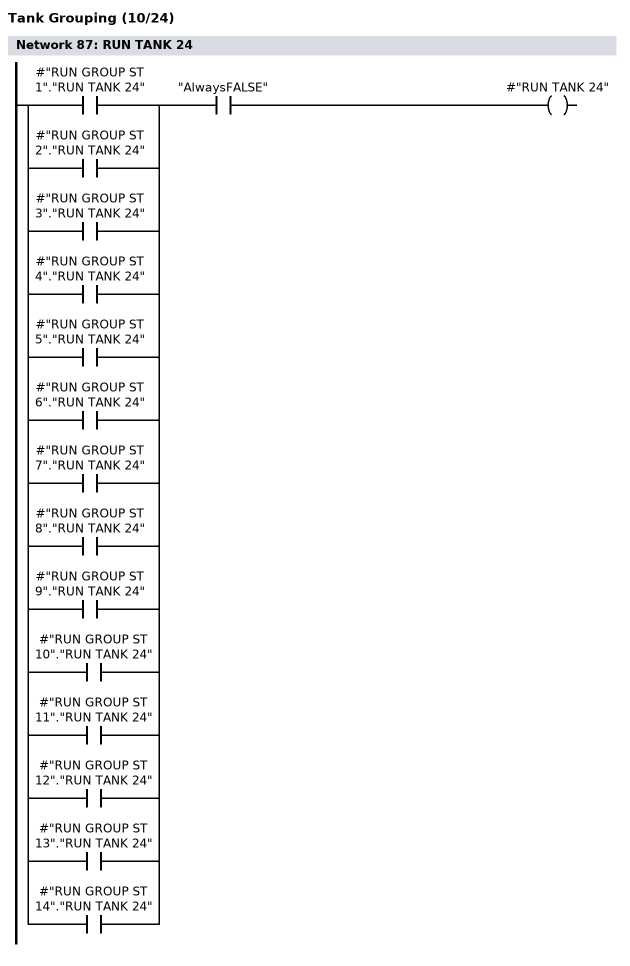
   RUNG wire#powerrail
      Contact( #"RUN GROUP ST 1"."RUN TANK 24" )
      wire#w1
      Contact( "AlwaysFALSE" )
      Coil( #"RUN TANK 24" )
   END_RUNG
   RUNG wire#powerrail
      Contact( #"RUN GROUP ST 2"."RUN TANK 24" )
   END_RUNG wire#w1
   RUNG wire#powerrail
      Contact( #"RUN GROUP ST 3"."RUN TANK 24" )
   END_RUNG wire#w1
   RUNG wire#powerrail
      Contact( #"RUN GROUP ST 4"."RUN TANK 24" )
   END_RUNG wire#w1
   RUNG wire#powerrail
      Contact( #"RUN GROUP ST 5"."RUN TANK 24" )
   END_RUNG wire#w1
   RUNG wire#powerrail
      Contact( #"RUN GROUP ST 6"."RUN TANK 24" )
   END_RUNG wire#w1
   RUNG wire#powerrail
      Contact( #"RUN GROUP ST 7"."RUN TANK 24" )
   END_RUNG wire#w1
   RUNG wire#powerrail
      Contact( #"RUN GROUP ST 8"."RUN TANK 24" )
   END_RUNG wire#w1
   RUNG wire#powerrail
      Contact( #"RUN GROUP ST 9"."RUN TANK 24" )
   END_RUNG wire#w1
   RUNG wire#powerrail
      Contact( #"RUN GROUP ST 10"."RUN TANK 24" )
   END_RUNG wire#w1
   RUNG wire#powerrail
      Contact( #"RUN GROUP ST 11"."RUN TANK 24" )
   END_RUNG wire#w1
   RUNG wire#powerrail
      Contact( #"RUN GROUP ST 12"."RUN TANK 24" )
   END_RUNG wire#w1
   RUNG wire#powerrail
      Contact( #"RUN GROUP ST 13"."RUN TANK 24" )
   END_RUNG wire#w1
   RUNG wire#powerrail
      Contact( #"RUN GROUP ST 14"."RUN TANK 24" )
   END_RUNG wire#w1
   // the same network as SCL:
   #"RUN TANK 24" := (#"RUN GROUP ST 1"."RUN TANK 24" OR #"RUN GROUP ST 2"."RUN TANK 24" OR #"RUN GROUP ST 3"."RUN TANK 24" OR #"RUN GROUP ST 4"."RUN TANK 24" OR #"RUN GROUP ST 5"."RUN TANK 24" OR #"RUN GROUP ST 6"."RUN TANK 24" OR #"RUN GROUP ST 7"."RUN TANK 24" OR #"RUN GROUP ST 8"."RUN TANK 24" OR #"RUN GROUP ST 9"."RUN TANK 24" OR #"RUN GROUP ST 10"."RUN TANK 24" OR #"RUN GROUP ST 11"."RUN TANK 24" OR #"RUN GROUP ST 12"."RUN TANK 24" OR #"RUN GROUP ST 13"."RUN TANK 24" OR #"RUN GROUP ST 14"."RUN TANK 24") AND "AlwaysFALSE";
END_REGION

REGION Network 89: Tank Selected Group 1
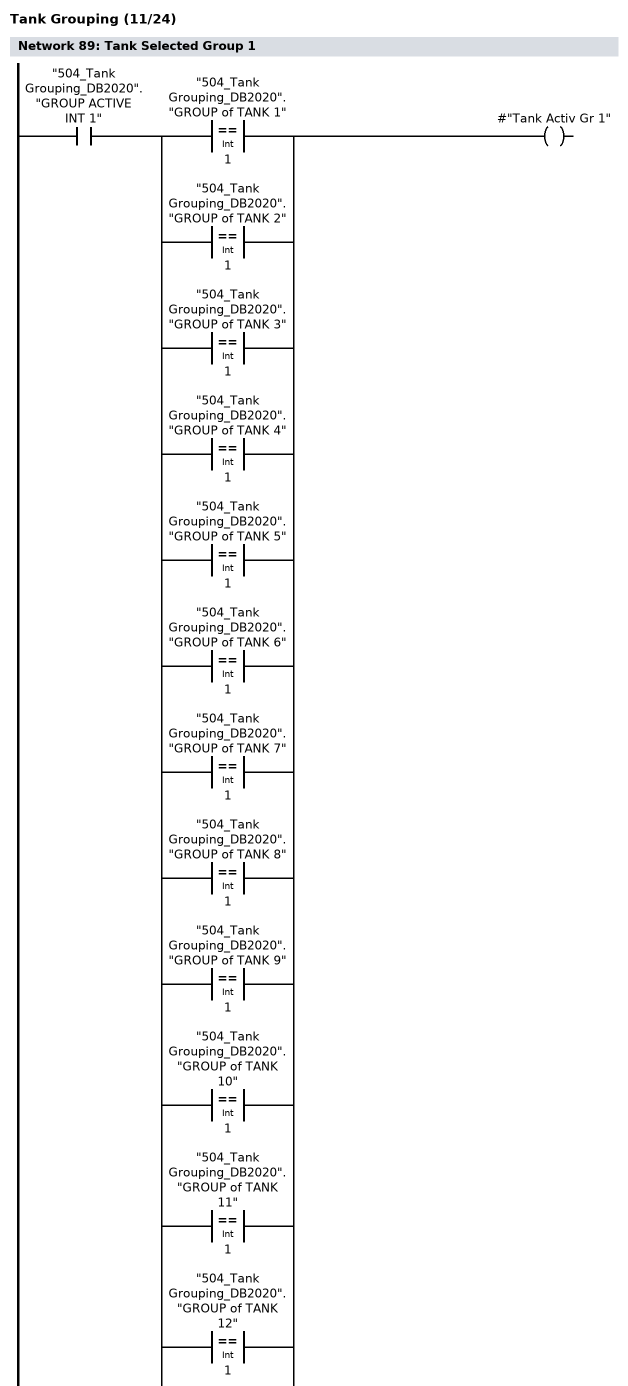
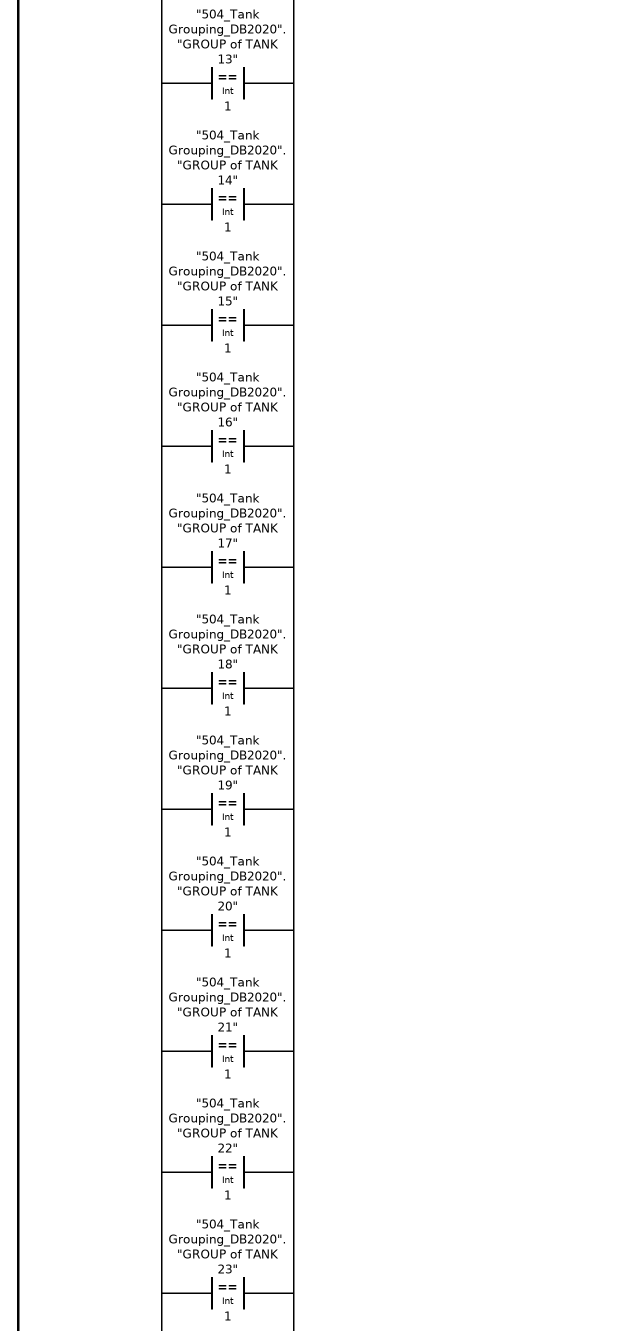
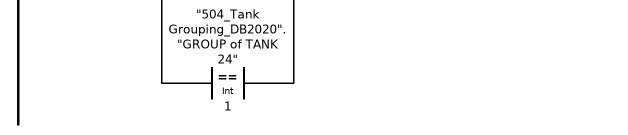
   RUNG wire#powerrail
      Contact( "504_Tank Grouping_DB2020"."GROUP ACTIVE INT 1" )
      wire#w1
      { S7_Templates := "SrcType := Int" } EQ_Contact(in1 := "504_Tank Grouping_DB2020"."GROUP of TANK 1", in2 := 1)
      wire#w2
      Coil( #"Tank Activ Gr 1" )
   END_RUNG
   RUNG wire#w1
      { S7_Templates := "SrcType := Int" } EQ_Contact(in1 := "504_Tank Grouping_DB2020"."GROUP of TANK 2", in2 := 1)
   END_RUNG wire#w2
   RUNG wire#w1
      { S7_Templates := "SrcType := Int" } EQ_Contact(in1 := "504_Tank Grouping_DB2020"."GROUP of TANK 3", in2 := 1)
   END_RUNG wire#w2
   RUNG wire#w1
      { S7_Templates := "SrcType := Int" } EQ_Contact(in1 := "504_Tank Grouping_DB2020"."GROUP of TANK 4", in2 := 1)
   END_RUNG wire#w2
   RUNG wire#w1
      { S7_Templates := "SrcType := Int" } EQ_Contact(in1 := "504_Tank Grouping_DB2020"."GROUP of TANK 5", in2 := 1)
   END_RUNG wire#w2
   RUNG wire#w1
      { S7_Templates := "SrcType := Int" } EQ_Contact(in1 := "504_Tank Grouping_DB2020"."GROUP of TANK 6", in2 := 1)
   END_RUNG wire#w2
   RUNG wire#w1
      { S7_Templates := "SrcType := Int" } EQ_Contact(in1 := "504_Tank Grouping_DB2020"."GROUP of TANK 7", in2 := 1)
   END_RUNG wire#w2
   RUNG wire#w1
      { S7_Templates := "SrcType := Int" } EQ_Contact(in1 := "504_Tank Grouping_DB2020"."GROUP of TANK 8", in2 := 1)
   END_RUNG wire#w2
   RUNG wire#w1
      { S7_Templates := "SrcType := Int" } EQ_Contact(in1 := "504_Tank Grouping_DB2020"."GROUP of TANK 9", in2 := 1)
   END_RUNG wire#w2
   RUNG wire#w1
      { S7_Templates := "SrcType := Int" } EQ_Contact(in1 := "504_Tank Grouping_DB2020"."GROUP of TANK 10", in2 := 1)
   END_RUNG wire#w2
   RUNG wire#w1
      { S7_Templates := "SrcType := Int" } EQ_Contact(in1 := "504_Tank Grouping_DB2020"."GROUP of TANK 11", in2 := 1)
   END_RUNG wire#w2
   RUNG wire#w1
      { S7_Templates := "SrcType := Int" } EQ_Contact(in1 := "504_Tank Grouping_DB2020"."GROUP of TANK 12", in2 := 1)
   END_RUNG wire#w2
   RUNG wire#w1
      { S7_Templates := "SrcType := Int" } EQ_Contact(in1 := "504_Tank Grouping_DB2020"."GROUP of TANK 13", in2 := 1)
   END_RUNG wire#w2
   RUNG wire#w1
      { S7_Templates := "SrcType := Int" } EQ_Contact(in1 := "504_Tank Grouping_DB2020"."GROUP of TANK 14", in2 := 1)
   END_RUNG wire#w2
   RUNG wire#w1
      { S7_Templates := "SrcType := Int" } EQ_Contact(in1 := "504_Tank Grouping_DB2020"."GROUP of TANK 15", in2 := 1)
   END_RUNG wire#w2
   RUNG wire#w1
      { S7_Templates := "SrcType := Int" } EQ_Contact(in1 := "504_Tank Grouping_DB2020"."GROUP of TANK 16", in2 := 1)
   END_RUNG wire#w2
   RUNG wire#w1
      { S7_Templates := "SrcType := Int" } EQ_Contact(in1 := "504_Tank Grouping_DB2020"."GROUP of TANK 17", in2 := 1)
   END_RUNG wire#w2
   RUNG wire#w1
      { S7_Templates := "SrcType := Int" } EQ_Contact(in1 := "504_Tank Grouping_DB2020"."GROUP of TANK 18", in2 := 1)
   END_RUNG wire#w2
   RUNG wire#w1
      { S7_Templates := "SrcType := Int" } EQ_Contact(in1 := "504_Tank Grouping_DB2020"."GROUP of TANK 19", in2 := 1)
   END_RUNG wire#w2
   RUNG wire#w1
      { S7_Templates := "SrcType := Int" } EQ_Contact(in1 := "504_Tank Grouping_DB2020"."GROUP of TANK 20", in2 := 1)
   END_RUNG wire#w2
   RUNG wire#w1
      { S7_Templates := "SrcType := Int" } EQ_Contact(in1 := "504_Tank Grouping_DB2020"."GROUP of TANK 21", in2 := 1)
   END_RUNG wire#w2
   RUNG wire#w1
      { S7_Templates := "SrcType := Int" } EQ_Contact(in1 := "504_Tank Grouping_DB2020"."GROUP of TANK 22", in2 := 1)
   END_RUNG wire#w2
   RUNG wire#w1
      { S7_Templates := "SrcType := Int" } EQ_Contact(in1 := "504_Tank Grouping_DB2020"."GROUP of TANK 23", in2 := 1)
   END_RUNG wire#w2
   RUNG wire#w1
      { S7_Templates := "SrcType := Int" } EQ_Contact(in1 := "504_Tank Grouping_DB2020"."GROUP of TANK 24", in2 := 1)
   END_RUNG wire#w2
   // the same network as SCL:
   #"Tank Activ Gr 1" := "504_Tank Grouping_DB2020"."GROUP ACTIVE INT 1" AND (("504_Tank Grouping_DB2020"."GROUP of TANK 1" = 1) OR ("504_Tank Grouping_DB2020"."GROUP of TANK 2" = 1) OR ("504_Tank Grouping_DB2020"."GROUP of TANK 3" = 1) OR ("504_Tank Grouping_DB2020"."GROUP of TANK 4" = 1) OR ("504_Tank Grouping_DB2020"."GROUP of TANK 5" = 1) OR ("504_Tank Grouping_DB2020"."GROUP of TANK 6" = 1) OR ("504_Tank Grouping_DB2020"."GROUP of TANK 7" = 1) OR ("504_Tank Grouping_DB2020"."GROUP of TANK 8" = 1) OR ("504_Tank Grouping_DB2020"."GROUP of TANK 9" = 1) OR ("504_Tank Grouping_DB2020"."GROUP of TANK 10" = 1) OR ("504_Tank Grouping_DB2020"."GROUP of TANK 11" = 1) OR ("504_Tank Grouping_DB2020"."GROUP of TANK 12" = 1) OR ("504_Tank Grouping_DB2020"."GROUP of TANK 13" = 1) OR ("504_Tank Grouping_DB2020"."GROUP of TANK 14" = 1) OR ("504_Tank Grouping_DB2020"."GROUP of TANK 15" = 1) OR ("504_Tank Grouping_DB2020"."GROUP of TANK 16" = 1) OR ("504_Tank Grouping_DB2020"."GROUP of TANK 17" = 1) OR ("504_Tank Grouping_DB2020"."GROUP of TANK 18" = 1) OR ("504_Tank Grouping_DB2020"."GROUP of TANK 19" = 1) OR ("504_Tank Grouping_DB2020"."GROUP of TANK 20" = 1) OR ("504_Tank Grouping_DB2020"."GROUP of TANK 21" = 1) OR ("504_Tank Grouping_DB2020"."GROUP of TANK 22" = 1) OR ("504_Tank Grouping_DB2020"."GROUP of TANK 23" = 1) OR ("504_Tank Grouping_DB2020"."GROUP of TANK 24" = 1));
END_REGION

REGION Network 90: Tank Selected Group 2
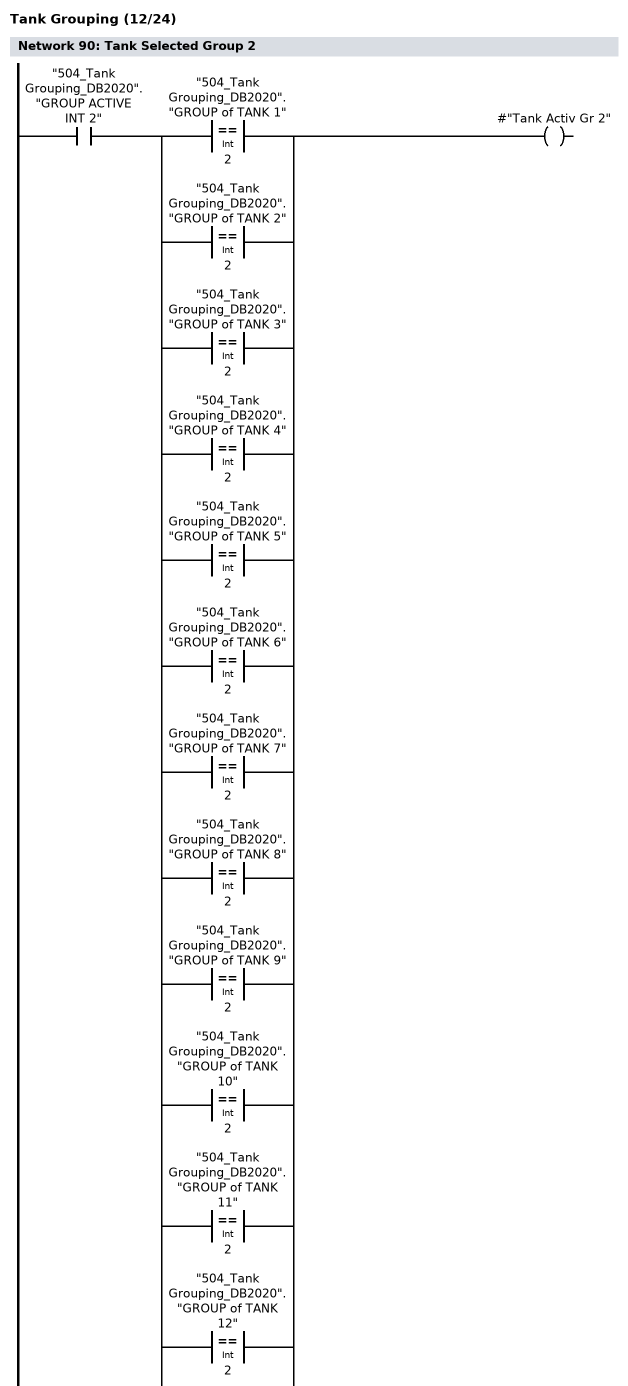
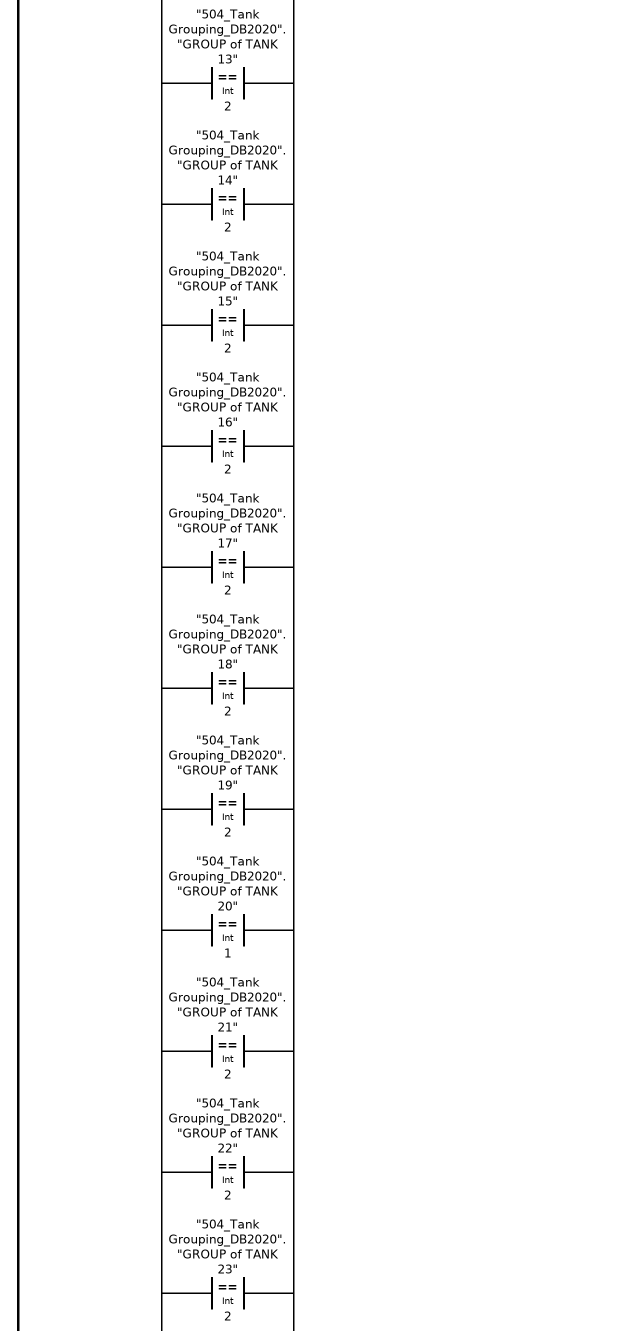
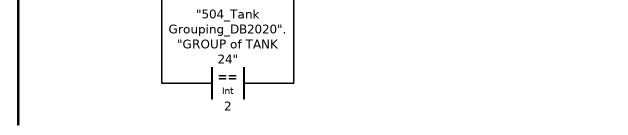
   RUNG wire#powerrail
      Contact( "504_Tank Grouping_DB2020"."GROUP ACTIVE INT 2" )
      wire#w1
      { S7_Templates := "SrcType := Int" } EQ_Contact(in1 := "504_Tank Grouping_DB2020"."GROUP of TANK 1", in2 := 2)
      wire#w2
      Coil( #"Tank Activ Gr 2" )
   END_RUNG
   RUNG wire#w1
      { S7_Templates := "SrcType := Int" } EQ_Contact(in1 := "504_Tank Grouping_DB2020"."GROUP of TANK 2", in2 := 2)
   END_RUNG wire#w2
   RUNG wire#w1
      { S7_Templates := "SrcType := Int" } EQ_Contact(in1 := "504_Tank Grouping_DB2020"."GROUP of TANK 3", in2 := 2)
   END_RUNG wire#w2
   RUNG wire#w1
      { S7_Templates := "SrcType := Int" } EQ_Contact(in1 := "504_Tank Grouping_DB2020"."GROUP of TANK 4", in2 := 2)
   END_RUNG wire#w2
   RUNG wire#w1
      { S7_Templates := "SrcType := Int" } EQ_Contact(in1 := "504_Tank Grouping_DB2020"."GROUP of TANK 5", in2 := 2)
   END_RUNG wire#w2
   RUNG wire#w1
      { S7_Templates := "SrcType := Int" } EQ_Contact(in1 := "504_Tank Grouping_DB2020"."GROUP of TANK 6", in2 := 2)
   END_RUNG wire#w2
   RUNG wire#w1
      { S7_Templates := "SrcType := Int" } EQ_Contact(in1 := "504_Tank Grouping_DB2020"."GROUP of TANK 7", in2 := 2)
   END_RUNG wire#w2
   RUNG wire#w1
      { S7_Templates := "SrcType := Int" } EQ_Contact(in1 := "504_Tank Grouping_DB2020"."GROUP of TANK 8", in2 := 2)
   END_RUNG wire#w2
   RUNG wire#w1
      { S7_Templates := "SrcType := Int" } EQ_Contact(in1 := "504_Tank Grouping_DB2020"."GROUP of TANK 9", in2 := 2)
   END_RUNG wire#w2
   RUNG wire#w1
      { S7_Templates := "SrcType := Int" } EQ_Contact(in1 := "504_Tank Grouping_DB2020"."GROUP of TANK 10", in2 := 2)
   END_RUNG wire#w2
   RUNG wire#w1
      { S7_Templates := "SrcType := Int" } EQ_Contact(in1 := "504_Tank Grouping_DB2020"."GROUP of TANK 11", in2 := 2)
   END_RUNG wire#w2
   RUNG wire#w1
      { S7_Templates := "SrcType := Int" } EQ_Contact(in1 := "504_Tank Grouping_DB2020"."GROUP of TANK 12", in2 := 2)
   END_RUNG wire#w2
   RUNG wire#w1
      { S7_Templates := "SrcType := Int" } EQ_Contact(in1 := "504_Tank Grouping_DB2020"."GROUP of TANK 13", in2 := 2)
   END_RUNG wire#w2
   RUNG wire#w1
      { S7_Templates := "SrcType := Int" } EQ_Contact(in1 := "504_Tank Grouping_DB2020"."GROUP of TANK 14", in2 := 2)
   END_RUNG wire#w2
   RUNG wire#w1
      { S7_Templates := "SrcType := Int" } EQ_Contact(in1 := "504_Tank Grouping_DB2020"."GROUP of TANK 15", in2 := 2)
   END_RUNG wire#w2
   RUNG wire#w1
      { S7_Templates := "SrcType := Int" } EQ_Contact(in1 := "504_Tank Grouping_DB2020"."GROUP of TANK 16", in2 := 2)
   END_RUNG wire#w2
   RUNG wire#w1
      { S7_Templates := "SrcType := Int" } EQ_Contact(in1 := "504_Tank Grouping_DB2020"."GROUP of TANK 17", in2 := 2)
   END_RUNG wire#w2
   RUNG wire#w1
      { S7_Templates := "SrcType := Int" } EQ_Contact(in1 := "504_Tank Grouping_DB2020"."GROUP of TANK 18", in2 := 2)
   END_RUNG wire#w2
   RUNG wire#w1
      { S7_Templates := "SrcType := Int" } EQ_Contact(in1 := "504_Tank Grouping_DB2020"."GROUP of TANK 19", in2 := 2)
   END_RUNG wire#w2
   RUNG wire#w1
      { S7_Templates := "SrcType := Int" } EQ_Contact(in1 := "504_Tank Grouping_DB2020"."GROUP of TANK 20", in2 := 1)
   END_RUNG wire#w2
   RUNG wire#w1
      { S7_Templates := "SrcType := Int" } EQ_Contact(in1 := "504_Tank Grouping_DB2020"."GROUP of TANK 21", in2 := 2)
   END_RUNG wire#w2
   RUNG wire#w1
      { S7_Templates := "SrcType := Int" } EQ_Contact(in1 := "504_Tank Grouping_DB2020"."GROUP of TANK 22", in2 := 2)
   END_RUNG wire#w2
   RUNG wire#w1
      { S7_Templates := "SrcType := Int" } EQ_Contact(in1 := "504_Tank Grouping_DB2020"."GROUP of TANK 23", in2 := 2)
   END_RUNG wire#w2
   RUNG wire#w1
      { S7_Templates := "SrcType := Int" } EQ_Contact(in1 := "504_Tank Grouping_DB2020"."GROUP of TANK 24", in2 := 2)
   END_RUNG wire#w2
   // the same network as SCL:
   #"Tank Activ Gr 2" := "504_Tank Grouping_DB2020"."GROUP ACTIVE INT 2" AND (("504_Tank Grouping_DB2020"."GROUP of TANK 1" = 2) OR ("504_Tank Grouping_DB2020"."GROUP of TANK 2" = 2) OR ("504_Tank Grouping_DB2020"."GROUP of TANK 3" = 2) OR ("504_Tank Grouping_DB2020"."GROUP of TANK 4" = 2) OR ("504_Tank Grouping_DB2020"."GROUP of TANK 5" = 2) OR ("504_Tank Grouping_DB2020"."GROUP of TANK 6" = 2) OR ("504_Tank Grouping_DB2020"."GROUP of TANK 7" = 2) OR ("504_Tank Grouping_DB2020"."GROUP of TANK 8" = 2) OR ("504_Tank Grouping_DB2020"."GROUP of TANK 9" = 2) OR ("504_Tank Grouping_DB2020"."GROUP of TANK 10" = 2) OR ("504_Tank Grouping_DB2020"."GROUP of TANK 11" = 2) OR ("504_Tank Grouping_DB2020"."GROUP of TANK 12" = 2) OR ("504_Tank Grouping_DB2020"."GROUP of TANK 13" = 2) OR ("504_Tank Grouping_DB2020"."GROUP of TANK 14" = 2) OR ("504_Tank Grouping_DB2020"."GROUP of TANK 15" = 2) OR ("504_Tank Grouping_DB2020"."GROUP of TANK 16" = 2) OR ("504_Tank Grouping_DB2020"."GROUP of TANK 17" = 2) OR ("504_Tank Grouping_DB2020"."GROUP of TANK 18" = 2) OR ("504_Tank Grouping_DB2020"."GROUP of TANK 19" = 2) OR ("504_Tank Grouping_DB2020"."GROUP of TANK 20" = 1) OR ("504_Tank Grouping_DB2020"."GROUP of TANK 21" = 2) OR ("504_Tank Grouping_DB2020"."GROUP of TANK 22" = 2) OR ("504_Tank Grouping_DB2020"."GROUP of TANK 23" = 2) OR ("504_Tank Grouping_DB2020"."GROUP of TANK 24" = 2));
END_REGION

REGION Network 91: Tank Selected Group 3
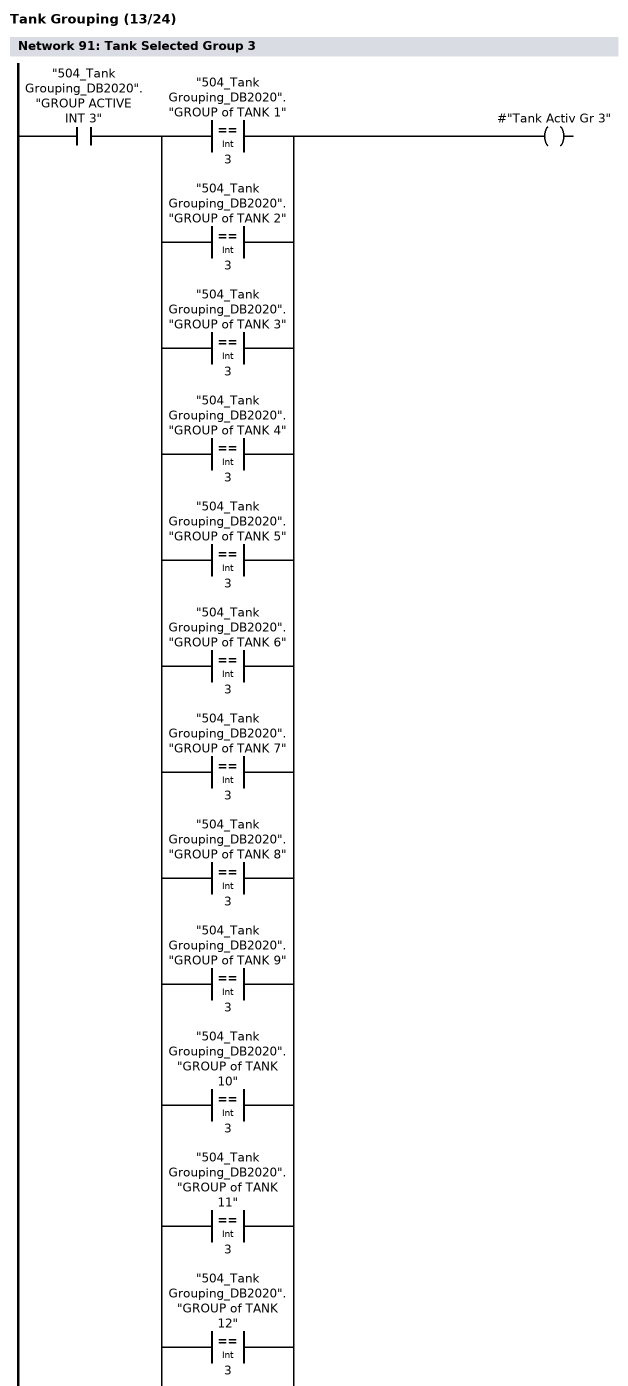
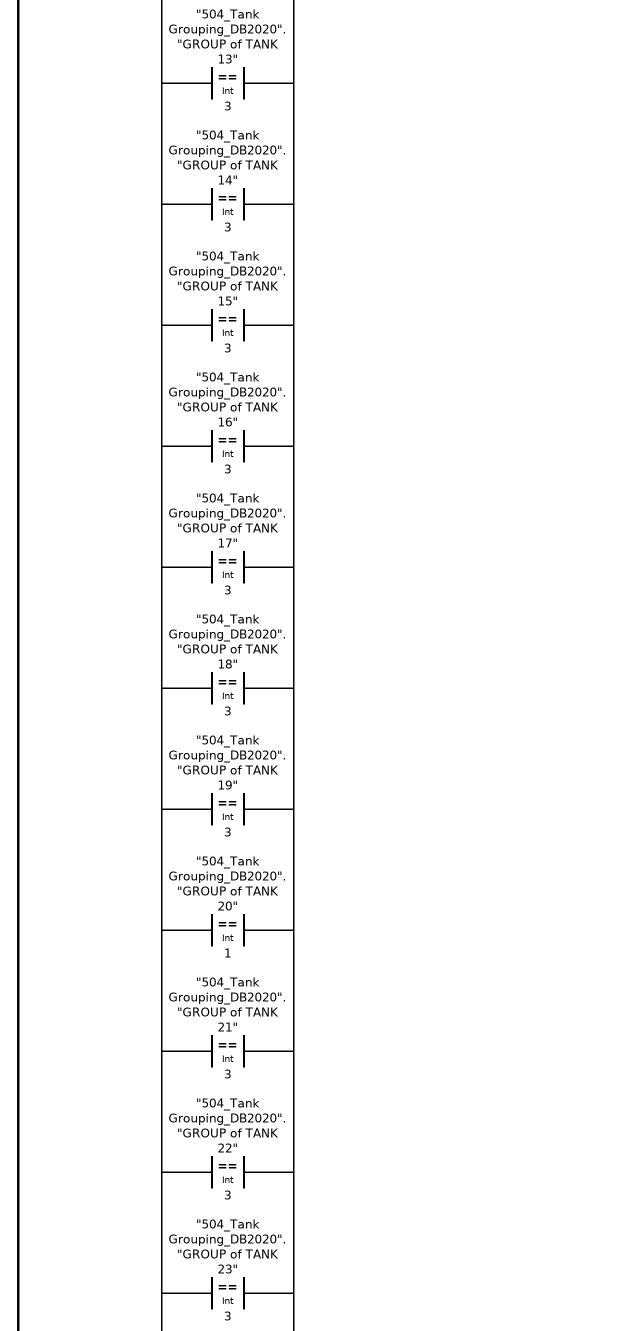
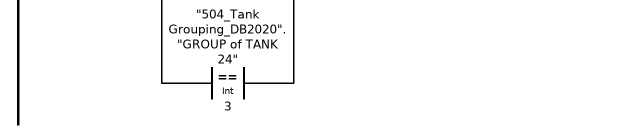
   RUNG wire#powerrail
      Contact( "504_Tank Grouping_DB2020"."GROUP ACTIVE INT 3" )
      wire#w1
      { S7_Templates := "SrcType := Int" } EQ_Contact(in1 := "504_Tank Grouping_DB2020"."GROUP of TANK 1", in2 := 3)
      wire#w2
      Coil( #"Tank Activ Gr 3" )
   END_RUNG
   RUNG wire#w1
      { S7_Templates := "SrcType := Int" } EQ_Contact(in1 := "504_Tank Grouping_DB2020"."GROUP of TANK 2", in2 := 3)
   END_RUNG wire#w2
   RUNG wire#w1
      { S7_Templates := "SrcType := Int" } EQ_Contact(in1 := "504_Tank Grouping_DB2020"."GROUP of TANK 3", in2 := 3)
   END_RUNG wire#w2
   RUNG wire#w1
      { S7_Templates := "SrcType := Int" } EQ_Contact(in1 := "504_Tank Grouping_DB2020"."GROUP of TANK 4", in2 := 3)
   END_RUNG wire#w2
   RUNG wire#w1
      { S7_Templates := "SrcType := Int" } EQ_Contact(in1 := "504_Tank Grouping_DB2020"."GROUP of TANK 5", in2 := 3)
   END_RUNG wire#w2
   RUNG wire#w1
      { S7_Templates := "SrcType := Int" } EQ_Contact(in1 := "504_Tank Grouping_DB2020"."GROUP of TANK 6", in2 := 3)
   END_RUNG wire#w2
   RUNG wire#w1
      { S7_Templates := "SrcType := Int" } EQ_Contact(in1 := "504_Tank Grouping_DB2020"."GROUP of TANK 7", in2 := 3)
   END_RUNG wire#w2
   RUNG wire#w1
      { S7_Templates := "SrcType := Int" } EQ_Contact(in1 := "504_Tank Grouping_DB2020"."GROUP of TANK 8", in2 := 3)
   END_RUNG wire#w2
   RUNG wire#w1
      { S7_Templates := "SrcType := Int" } EQ_Contact(in1 := "504_Tank Grouping_DB2020"."GROUP of TANK 9", in2 := 3)
   END_RUNG wire#w2
   RUNG wire#w1
      { S7_Templates := "SrcType := Int" } EQ_Contact(in1 := "504_Tank Grouping_DB2020"."GROUP of TANK 10", in2 := 3)
   END_RUNG wire#w2
   RUNG wire#w1
      { S7_Templates := "SrcType := Int" } EQ_Contact(in1 := "504_Tank Grouping_DB2020"."GROUP of TANK 11", in2 := 3)
   END_RUNG wire#w2
   RUNG wire#w1
      { S7_Templates := "SrcType := Int" } EQ_Contact(in1 := "504_Tank Grouping_DB2020"."GROUP of TANK 12", in2 := 3)
   END_RUNG wire#w2
   RUNG wire#w1
      { S7_Templates := "SrcType := Int" } EQ_Contact(in1 := "504_Tank Grouping_DB2020"."GROUP of TANK 13", in2 := 3)
   END_RUNG wire#w2
   RUNG wire#w1
      { S7_Templates := "SrcType := Int" } EQ_Contact(in1 := "504_Tank Grouping_DB2020"."GROUP of TANK 14", in2 := 3)
   END_RUNG wire#w2
   RUNG wire#w1
      { S7_Templates := "SrcType := Int" } EQ_Contact(in1 := "504_Tank Grouping_DB2020"."GROUP of TANK 15", in2 := 3)
   END_RUNG wire#w2
   RUNG wire#w1
      { S7_Templates := "SrcType := Int" } EQ_Contact(in1 := "504_Tank Grouping_DB2020"."GROUP of TANK 16", in2 := 3)
   END_RUNG wire#w2
   RUNG wire#w1
      { S7_Templates := "SrcType := Int" } EQ_Contact(in1 := "504_Tank Grouping_DB2020"."GROUP of TANK 17", in2 := 3)
   END_RUNG wire#w2
   RUNG wire#w1
      { S7_Templates := "SrcType := Int" } EQ_Contact(in1 := "504_Tank Grouping_DB2020"."GROUP of TANK 18", in2 := 3)
   END_RUNG wire#w2
   RUNG wire#w1
      { S7_Templates := "SrcType := Int" } EQ_Contact(in1 := "504_Tank Grouping_DB2020"."GROUP of TANK 19", in2 := 3)
   END_RUNG wire#w2
   RUNG wire#w1
      { S7_Templates := "SrcType := Int" } EQ_Contact(in1 := "504_Tank Grouping_DB2020"."GROUP of TANK 20", in2 := 1)
   END_RUNG wire#w2
   RUNG wire#w1
      { S7_Templates := "SrcType := Int" } EQ_Contact(in1 := "504_Tank Grouping_DB2020"."GROUP of TANK 21", in2 := 3)
   END_RUNG wire#w2
   RUNG wire#w1
      { S7_Templates := "SrcType := Int" } EQ_Contact(in1 := "504_Tank Grouping_DB2020"."GROUP of TANK 22", in2 := 3)
   END_RUNG wire#w2
   RUNG wire#w1
      { S7_Templates := "SrcType := Int" } EQ_Contact(in1 := "504_Tank Grouping_DB2020"."GROUP of TANK 23", in2 := 3)
   END_RUNG wire#w2
   RUNG wire#w1
      { S7_Templates := "SrcType := Int" } EQ_Contact(in1 := "504_Tank Grouping_DB2020"."GROUP of TANK 24", in2 := 3)
   END_RUNG wire#w2
   // the same network as SCL:
   #"Tank Activ Gr 3" := "504_Tank Grouping_DB2020"."GROUP ACTIVE INT 3" AND (("504_Tank Grouping_DB2020"."GROUP of TANK 1" = 3) OR ("504_Tank Grouping_DB2020"."GROUP of TANK 2" = 3) OR ("504_Tank Grouping_DB2020"."GROUP of TANK 3" = 3) OR ("504_Tank Grouping_DB2020"."GROUP of TANK 4" = 3) OR ("504_Tank Grouping_DB2020"."GROUP of TANK 5" = 3) OR ("504_Tank Grouping_DB2020"."GROUP of TANK 6" = 3) OR ("504_Tank Grouping_DB2020"."GROUP of TANK 7" = 3) OR ("504_Tank Grouping_DB2020"."GROUP of TANK 8" = 3) OR ("504_Tank Grouping_DB2020"."GROUP of TANK 9" = 3) OR ("504_Tank Grouping_DB2020"."GROUP of TANK 10" = 3) OR ("504_Tank Grouping_DB2020"."GROUP of TANK 11" = 3) OR ("504_Tank Grouping_DB2020"."GROUP of TANK 12" = 3) OR ("504_Tank Grouping_DB2020"."GROUP of TANK 13" = 3) OR ("504_Tank Grouping_DB2020"."GROUP of TANK 14" = 3) OR ("504_Tank Grouping_DB2020"."GROUP of TANK 15" = 3) OR ("504_Tank Grouping_DB2020"."GROUP of TANK 16" = 3) OR ("504_Tank Grouping_DB2020"."GROUP of TANK 17" = 3) OR ("504_Tank Grouping_DB2020"."GROUP of TANK 18" = 3) OR ("504_Tank Grouping_DB2020"."GROUP of TANK 19" = 3) OR ("504_Tank Grouping_DB2020"."GROUP of TANK 20" = 1) OR ("504_Tank Grouping_DB2020"."GROUP of TANK 21" = 3) OR ("504_Tank Grouping_DB2020"."GROUP of TANK 22" = 3) OR ("504_Tank Grouping_DB2020"."GROUP of TANK 23" = 3) OR ("504_Tank Grouping_DB2020"."GROUP of TANK 24" = 3));
END_REGION

REGION Network 92: Tank Selected Group 4
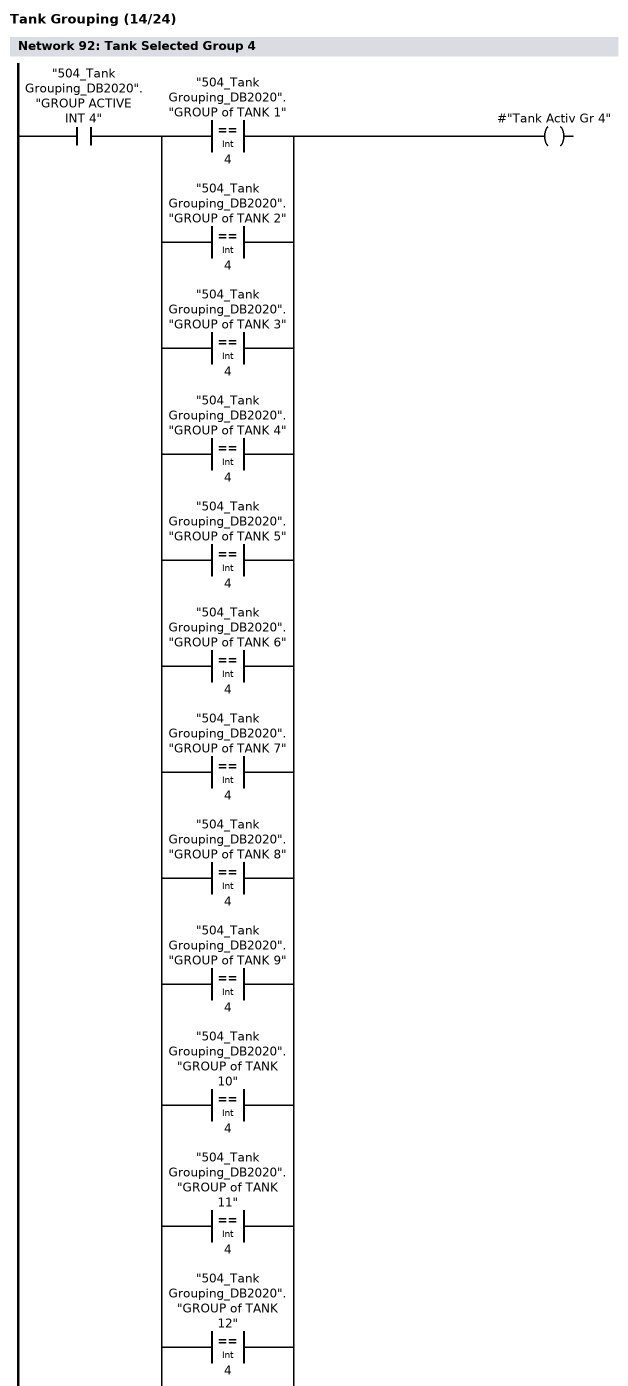
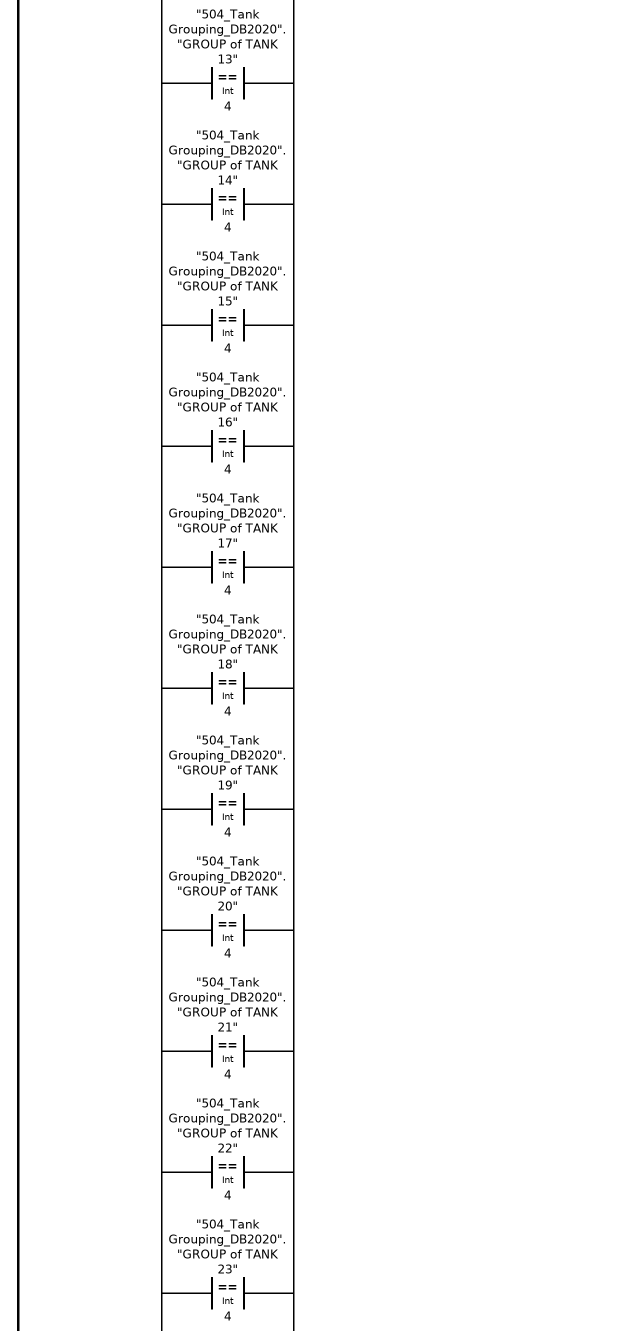
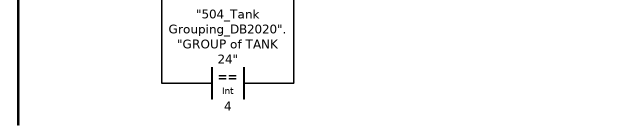
   RUNG wire#powerrail
      Contact( "504_Tank Grouping_DB2020"."GROUP ACTIVE INT 4" )
      wire#w1
      { S7_Templates := "SrcType := Int" } EQ_Contact(in1 := "504_Tank Grouping_DB2020"."GROUP of TANK 1", in2 := 4)
      wire#w2
      Coil( #"Tank Activ Gr 4" )
   END_RUNG
   RUNG wire#w1
      { S7_Templates := "SrcType := Int" } EQ_Contact(in1 := "504_Tank Grouping_DB2020"."GROUP of TANK 2", in2 := 4)
   END_RUNG wire#w2
   RUNG wire#w1
      { S7_Templates := "SrcType := Int" } EQ_Contact(in1 := "504_Tank Grouping_DB2020"."GROUP of TANK 3", in2 := 4)
   END_RUNG wire#w2
   RUNG wire#w1
      { S7_Templates := "SrcType := Int" } EQ_Contact(in1 := "504_Tank Grouping_DB2020"."GROUP of TANK 4", in2 := 4)
   END_RUNG wire#w2
   RUNG wire#w1
      { S7_Templates := "SrcType := Int" } EQ_Contact(in1 := "504_Tank Grouping_DB2020"."GROUP of TANK 5", in2 := 4)
   END_RUNG wire#w2
   RUNG wire#w1
      { S7_Templates := "SrcType := Int" } EQ_Contact(in1 := "504_Tank Grouping_DB2020"."GROUP of TANK 6", in2 := 4)
   END_RUNG wire#w2
   RUNG wire#w1
      { S7_Templates := "SrcType := Int" } EQ_Contact(in1 := "504_Tank Grouping_DB2020"."GROUP of TANK 7", in2 := 4)
   END_RUNG wire#w2
   RUNG wire#w1
      { S7_Templates := "SrcType := Int" } EQ_Contact(in1 := "504_Tank Grouping_DB2020"."GROUP of TANK 8", in2 := 4)
   END_RUNG wire#w2
   RUNG wire#w1
      { S7_Templates := "SrcType := Int" } EQ_Contact(in1 := "504_Tank Grouping_DB2020"."GROUP of TANK 9", in2 := 4)
   END_RUNG wire#w2
   RUNG wire#w1
      { S7_Templates := "SrcType := Int" } EQ_Contact(in1 := "504_Tank Grouping_DB2020"."GROUP of TANK 10", in2 := 4)
   END_RUNG wire#w2
   RUNG wire#w1
      { S7_Templates := "SrcType := Int" } EQ_Contact(in1 := "504_Tank Grouping_DB2020"."GROUP of TANK 11", in2 := 4)
   END_RUNG wire#w2
   RUNG wire#w1
      { S7_Templates := "SrcType := Int" } EQ_Contact(in1 := "504_Tank Grouping_DB2020"."GROUP of TANK 12", in2 := 4)
   END_RUNG wire#w2
   RUNG wire#w1
      { S7_Templates := "SrcType := Int" } EQ_Contact(in1 := "504_Tank Grouping_DB2020"."GROUP of TANK 13", in2 := 4)
   END_RUNG wire#w2
   RUNG wire#w1
      { S7_Templates := "SrcType := Int" } EQ_Contact(in1 := "504_Tank Grouping_DB2020"."GROUP of TANK 14", in2 := 4)
   END_RUNG wire#w2
   RUNG wire#w1
      { S7_Templates := "SrcType := Int" } EQ_Contact(in1 := "504_Tank Grouping_DB2020"."GROUP of TANK 15", in2 := 4)
   END_RUNG wire#w2
   RUNG wire#w1
      { S7_Templates := "SrcType := Int" } EQ_Contact(in1 := "504_Tank Grouping_DB2020"."GROUP of TANK 16", in2 := 4)
   END_RUNG wire#w2
   RUNG wire#w1
      { S7_Templates := "SrcType := Int" } EQ_Contact(in1 := "504_Tank Grouping_DB2020"."GROUP of TANK 17", in2 := 4)
   END_RUNG wire#w2
   RUNG wire#w1
      { S7_Templates := "SrcType := Int" } EQ_Contact(in1 := "504_Tank Grouping_DB2020"."GROUP of TANK 18", in2 := 4)
   END_RUNG wire#w2
   RUNG wire#w1
      { S7_Templates := "SrcType := Int" } EQ_Contact(in1 := "504_Tank Grouping_DB2020"."GROUP of TANK 19", in2 := 4)
   END_RUNG wire#w2
   RUNG wire#w1
      { S7_Templates := "SrcType := Int" } EQ_Contact(in1 := "504_Tank Grouping_DB2020"."GROUP of TANK 20", in2 := 4)
   END_RUNG wire#w2
   RUNG wire#w1
      { S7_Templates := "SrcType := Int" } EQ_Contact(in1 := "504_Tank Grouping_DB2020"."GROUP of TANK 21", in2 := 4)
   END_RUNG wire#w2
   RUNG wire#w1
      { S7_Templates := "SrcType := Int" } EQ_Contact(in1 := "504_Tank Grouping_DB2020"."GROUP of TANK 22", in2 := 4)
   END_RUNG wire#w2
   RUNG wire#w1
      { S7_Templates := "SrcType := Int" } EQ_Contact(in1 := "504_Tank Grouping_DB2020"."GROUP of TANK 23", in2 := 4)
   END_RUNG wire#w2
   RUNG wire#w1
      { S7_Templates := "SrcType := Int" } EQ_Contact(in1 := "504_Tank Grouping_DB2020"."GROUP of TANK 24", in2 := 4)
   END_RUNG wire#w2
   // the same network as SCL:
   #"Tank Activ Gr 4" := "504_Tank Grouping_DB2020"."GROUP ACTIVE INT 4" AND (("504_Tank Grouping_DB2020"."GROUP of TANK 1" = 4) OR ("504_Tank Grouping_DB2020"."GROUP of TANK 2" = 4) OR ("504_Tank Grouping_DB2020"."GROUP of TANK 3" = 4) OR ("504_Tank Grouping_DB2020"."GROUP of TANK 4" = 4) OR ("504_Tank Grouping_DB2020"."GROUP of TANK 5" = 4) OR ("504_Tank Grouping_DB2020"."GROUP of TANK 6" = 4) OR ("504_Tank Grouping_DB2020"."GROUP of TANK 7" = 4) OR ("504_Tank Grouping_DB2020"."GROUP of TANK 8" = 4) OR ("504_Tank Grouping_DB2020"."GROUP of TANK 9" = 4) OR ("504_Tank Grouping_DB2020"."GROUP of TANK 10" = 4) OR ("504_Tank Grouping_DB2020"."GROUP of TANK 11" = 4) OR ("504_Tank Grouping_DB2020"."GROUP of TANK 12" = 4) OR ("504_Tank Grouping_DB2020"."GROUP of TANK 13" = 4) OR ("504_Tank Grouping_DB2020"."GROUP of TANK 14" = 4) OR ("504_Tank Grouping_DB2020"."GROUP of TANK 15" = 4) OR ("504_Tank Grouping_DB2020"."GROUP of TANK 16" = 4) OR ("504_Tank Grouping_DB2020"."GROUP of TANK 17" = 4) OR ("504_Tank Grouping_DB2020"."GROUP of TANK 18" = 4) OR ("504_Tank Grouping_DB2020"."GROUP of TANK 19" = 4) OR ("504_Tank Grouping_DB2020"."GROUP of TANK 20" = 4) OR ("504_Tank Grouping_DB2020"."GROUP of TANK 21" = 4) OR ("504_Tank Grouping_DB2020"."GROUP of TANK 22" = 4) OR ("504_Tank Grouping_DB2020"."GROUP of TANK 23" = 4) OR ("504_Tank Grouping_DB2020"."GROUP of TANK 24" = 4));
END_REGION

REGION Network 93: Tank Selected Group 5
